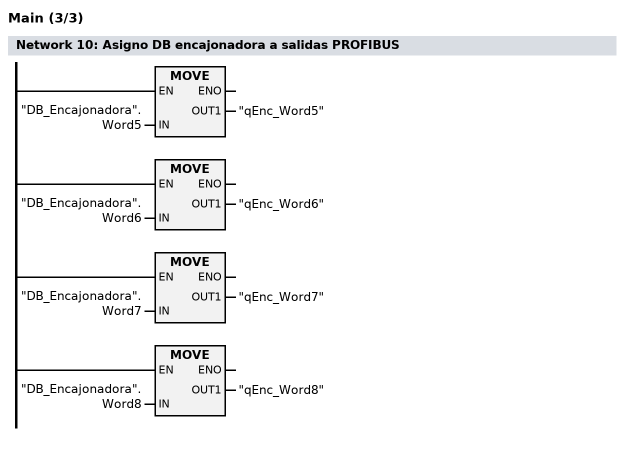
   RUNG wire#powerrail
      Move(in := "DB_Encajonadora".Word5, out1 => "qEnc_Word5")
   END_RUNG
   RUNG wire#powerrail
      Move(in := "DB_Encajonadora".Word6, out1 => "qEnc_Word6")
   END_RUNG
   RUNG wire#powerrail
      Move(in := "DB_Encajonadora".Word7, out1 => "qEnc_Word7")
   END_RUNG
   RUNG wire#powerrail
      Move(in := "DB_Encajonadora".Word8, out1 => "qEnc_Word8")
   END_RUNG
   // the same network as SCL:
   "qEnc_Word5" := "DB_Encajonadora".Word5;
   "qEnc_Word6" := "DB_Encajonadora".Word6;
   "qEnc_Word7" := "DB_Encajonadora".Word7;
   "qEnc_Word8" := "DB_Encajonadora".Word8;
END_REGION
END_ORGANIZATION_BLOCK

ORGANIZATION_BLOCK "Cyclic interrupt"   // OB30, LAD, CyclicInterrupt
{ S7_Optimized_Access := 'TRUE' }
VERSION : 0.1
   VAR_INPUT
      Initial_Call : Bool;   // Initial call of this OB
      Event_Count : Int;   // Events discarded
   END_VAR
BEGIN

REGION Network 1: Move
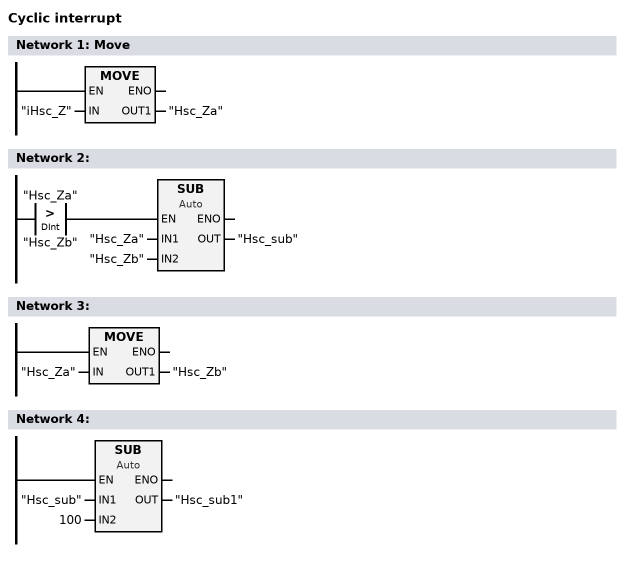
   RUNG wire#powerrail
      Move(in := "iHsc_Z", out1 => "Hsc_Za")
   END_RUNG
   // the same network as SCL:
   "Hsc_Za" := "iHsc_Z";
END_REGION

REGION Network 2
   RUNG wire#powerrail
      { S7_Templates := "SrcType := DInt" } GT_Contact(in1 := "Hsc_Za", in2 := "Hsc_Zb")
      Sub(in1 := "Hsc_Za", in2 := "Hsc_Zb", out => "Hsc_sub")
   END_RUNG
   // the same network as SCL:
   IF "Hsc_Za" > "Hsc_Zb" THEN "Hsc_sub" := "Hsc_Za" - "Hsc_Zb"; END_IF;
END_REGION

REGION Network 3
   RUNG wire#powerrail
      Move(in := "Hsc_Za", out1 => "Hsc_Zb")
   END_RUNG
   // the same network as SCL:
   "Hsc_Zb" := "Hsc_Za";
END_REGION

REGION Network 4
   RUNG wire#powerrail
      Sub(in1 := "Hsc_sub", in2 := 100, out => "Hsc_sub1")
   END_RUNG
   // the same network as SCL:
   "Hsc_sub1" := "Hsc_sub" - 100;
END_REGION
END_ORGANIZATION_BLOCK

// folder: ESTANDAR

FUNCTION_BLOCK "Motor M&CM"   // FB2, LAD
TITLE = Motor Marcha & Contra-Marcha
{ S7_Optimized_Access := 'TRUE' }
VERSION : 0.1
   VAR_INPUT
      iOrdMar_Dir : Bool;
      iOrdMar_Rev : Bool;
      iConfMar_Dir : Bool;
      iConfMar_Rev : Bool;
      iGMT : Bool;
      iTConf_Warn : Time;
      iTConf_Fall : Time;
      iTRearranque : Time;
   END_VAR
   VAR_OUTPUT
      oMar_Dir : Bool;
      oMar_Rev : Bool;
      oWarning_CTC_Dir : Bool;
      oWarning_CTC_Rev : Bool;
      oFall_CTC_Dir : Bool;
      oFall_CTC_Rev : Bool;
      oFall_GMT : Bool;
   END_VAR
   VAR
      IEC_Timer_0_Instance : IEC_TIMER;
      IEC_Timer_0_Instance_1 : IEC_TIMER;
      IEC_Timer_0_Instance_2 : IEC_TIMER;
      IEC_Timer_0_Instance_3 : IEC_TIMER;
      IEC_Timer_0_Instance_4 : IEC_TIMER;
      MarDir_Aux : Bool;
      MarRev_Aux : Bool;
   END_VAR
   VAR_TEMP
      Fall_GMT_Aux : Bool;
      Fall_CTC_Dir_Aux : Bool;
      Fall_CTC_Rev_Aux : Bool;
      Habil_Mov : Bool;
   END_VAR
   VAR_TEMP   // added for the SCL form of the ladder/FBD networks
      _w1 : Bool;
   END_VAR
BEGIN

REGION Network 1: Falla Guardamotor
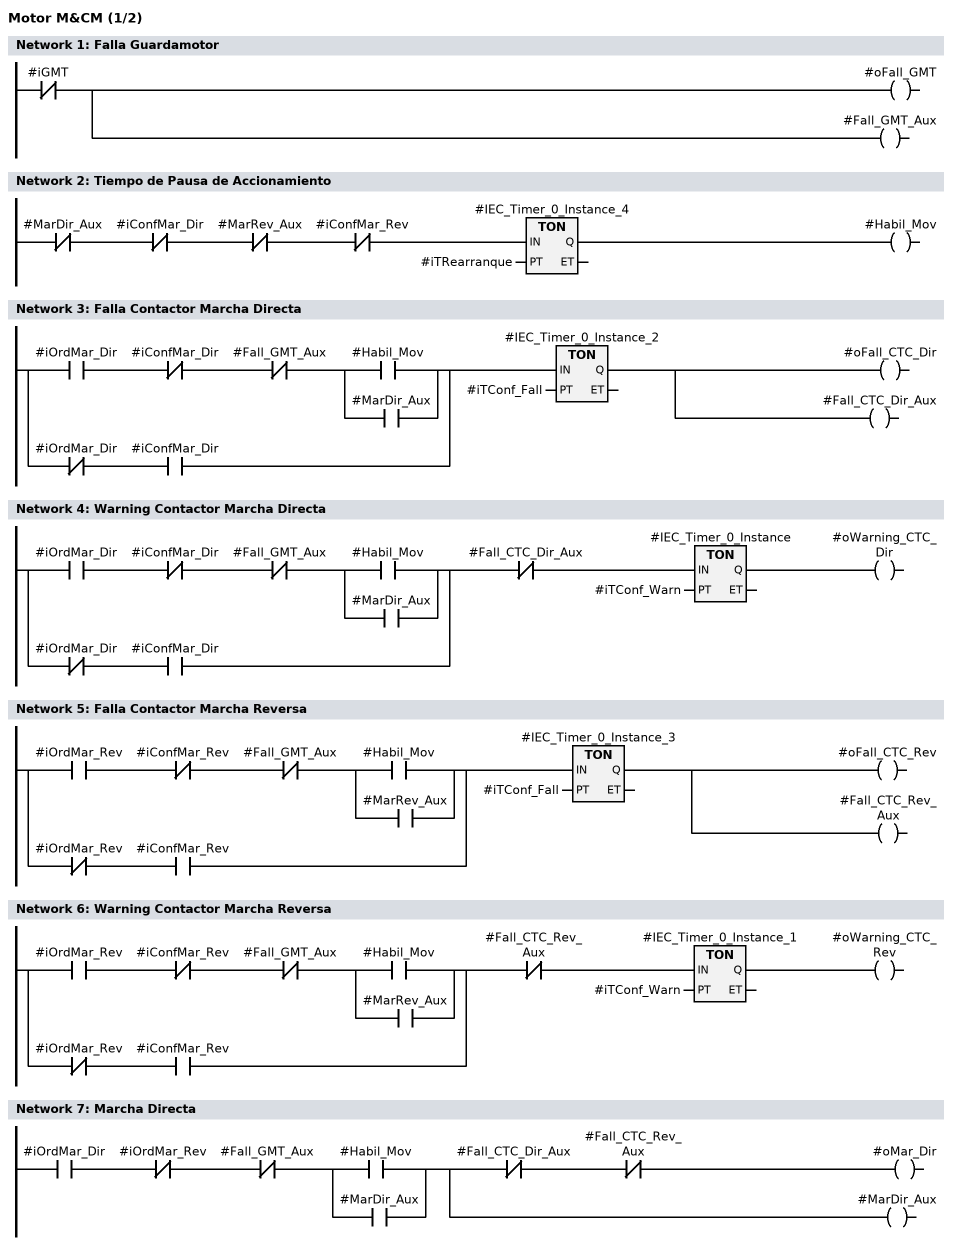
   RUNG wire#powerrail
      I_Contact( #iGMT )
      wire#w1
      Coil( #oFall_GMT )
   END_RUNG
   RUNG wire#w1
      Coil( #Fall_GMT_Aux )
   END_RUNG
   // the same network as SCL:
   #oFall_GMT := NOT #iGMT;
   #Fall_GMT_Aux := NOT #iGMT;
END_REGION

REGION Network 2: Tiempo de Pausa de Accionamiento
   #IEC_Timer_0_Instance_4.TON(IN := NOT #MarDir_Aux AND NOT #iConfMar_Dir AND NOT #MarRev_Aux AND NOT #iConfMar_Rev,
                           PT := #iTRearranque);
   #Habil_Mov := #IEC_Timer_0_Instance_4.Q;
END_REGION

REGION Network 3: Falla Contactor Marcha Directa
   #IEC_Timer_0_Instance_2.TON(IN := (#iOrdMar_Dir AND NOT #iConfMar_Dir AND NOT #Fall_GMT_Aux AND (#Habil_Mov OR #MarDir_Aux)) OR (NOT #iOrdMar_Dir AND #iConfMar_Dir),
                           PT := #iTConf_Fall);
   #oFall_CTC_Dir := #IEC_Timer_0_Instance_2.Q;
   #Fall_CTC_Dir_Aux := #IEC_Timer_0_Instance_2.Q;
END_REGION

REGION Network 4: Warning Contactor Marcha Directa
   #IEC_Timer_0_Instance.TON(IN := ((#iOrdMar_Dir AND NOT #iConfMar_Dir AND NOT #Fall_GMT_Aux AND (#Habil_Mov OR #MarDir_Aux)) OR (NOT #iOrdMar_Dir AND #iConfMar_Dir)) AND NOT #Fall_CTC_Dir_Aux,
                           PT := #iTConf_Warn);
   #oWarning_CTC_Dir := #IEC_Timer_0_Instance.Q;
END_REGION

REGION Network 5: Falla Contactor Marcha Reversa
   #IEC_Timer_0_Instance_3.TON(IN := (#iOrdMar_Rev AND NOT #iConfMar_Rev AND NOT #Fall_GMT_Aux AND (#Habil_Mov OR #MarRev_Aux)) OR (NOT #iOrdMar_Rev AND #iConfMar_Rev),
                           PT := #iTConf_Fall);
   #oFall_CTC_Rev := #IEC_Timer_0_Instance_3.Q;
   #Fall_CTC_Rev_Aux := #IEC_Timer_0_Instance_3.Q;
END_REGION

REGION Network 6: Warning Contactor Marcha Reversa
   #IEC_Timer_0_Instance_1.TON(IN := ((#iOrdMar_Rev AND NOT #iConfMar_Rev AND NOT #Fall_GMT_Aux AND (#Habil_Mov OR #MarRev_Aux)) OR (NOT #iOrdMar_Rev AND #iConfMar_Rev)) AND NOT #Fall_CTC_Rev_Aux,
                           PT := #iTConf_Warn);
   #oWarning_CTC_Rev := #IEC_Timer_0_Instance_1.Q;
END_REGION

REGION Network 7: Marcha Directa
   RUNG wire#powerrail
      Contact( #iOrdMar_Dir )
      I_Contact( #iOrdMar_Rev )
      I_Contact( #Fall_GMT_Aux )
      wire#w1
      Contact( #Habil_Mov )
      wire#w2
      I_Contact( #Fall_CTC_Dir_Aux )
      I_Contact( #Fall_CTC_Rev_Aux )
      Coil( #oMar_Dir )
   END_RUNG
   RUNG wire#w1
      Contact( #MarDir_Aux )
   END_RUNG wire#w2
   RUNG wire#w2
      Coil( #MarDir_Aux )
   END_RUNG
   // the same network as SCL:
   #_w1 := #iOrdMar_Dir AND NOT #iOrdMar_Rev AND NOT #Fall_GMT_Aux AND (#Habil_Mov OR #MarDir_Aux);
   #oMar_Dir := #_w1 AND NOT #Fall_CTC_Dir_Aux AND NOT #Fall_CTC_Rev_Aux;
   #MarDir_Aux := #_w1;
END_REGION

REGION Network 8: Marcha Reversa
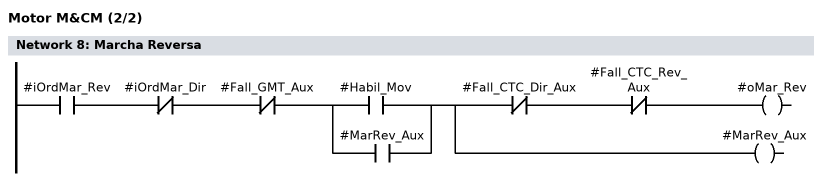
   RUNG wire#powerrail
      Contact( #iOrdMar_Rev )
      I_Contact( #iOrdMar_Dir )
      I_Contact( #Fall_GMT_Aux )
      wire#w1
      Contact( #Habil_Mov )
      wire#w2
      I_Contact( #Fall_CTC_Dir_Aux )
      I_Contact( #Fall_CTC_Rev_Aux )
      Coil( #oMar_Rev )
   END_RUNG
   RUNG wire#w1
      Contact( #MarRev_Aux )
   END_RUNG wire#w2
   RUNG wire#w2
      Coil( #MarRev_Aux )
   END_RUNG
   // the same network as SCL:
   #_w1 := #iOrdMar_Rev AND NOT #iOrdMar_Dir AND NOT #Fall_GMT_Aux AND (#Habil_Mov OR #MarRev_Aux);
   #oMar_Rev := #_w1 AND NOT #Fall_CTC_Dir_Aux AND NOT #Fall_CTC_Rev_Aux;
   #MarRev_Aux := #_w1;
END_REGION
END_FUNCTION_BLOCK

FUNCTION_BLOCK "FB_VAR_MOT"   // FB4, LAD
{ S7_Optimized_Access := 'FALSE' }
VERSION : 0.1
   VAR_INPUT
      "CMD Mar Dir" : Bool;   // Comando Marcha Directa
      "CMD Mar Rev" : Bool;   // Comando Marcha Reversa
      "HAB  Mar" : Bool;   // Habilita Marcha
      "SP Vel" : Real;   // Setpoint de Velocidad
      Reset : Bool;   // Comando resetear falla
      Fault : Bool;   // Indica variador en falla
      Ready : Bool;   // Indica variador Ready
      Ton_Freno : Time := T#400ms;
      Ton_Mar : Time := T#100ms;
      Tof_Freno : Time := T#100ms;
      Tof_Mar : Time := T#200ms;
   END_VAR
   VAR_OUTPUT
      Marcha : Bool;   // Orden de marcha a variador
      "Inv Giro" : Bool;   // Orden de invertir sentido de giro a variador
      "Reset Fault" : Bool;   // Reset Fault a variador
      Velocidad : Word;   // Referencia de Velocidad a variador
      Freno : Bool;   // Apertura de Freno
      Falla : Bool;   // Indica falla del variador
      Warning : Bool;   // Indica variador no Ready
   END_VAR
   VAR
      IEC_Timer_Freno : TON_TIME;
      IEC_Timer_Motor : TON_TIME;
      IEC_Timer_Reset : TOF_TIME;
      "_CMD Marcha Dir" : Bool;
      "_CMD Marcha Rev" : Bool;
      _CMD_AbrirFreno : Bool;
      IEC_Timer_0_Instance : TON_TIME;
      IEC_Timer_0_Instance_1 : TOF_TIME;
      IEC_Timer_0_Instance_2 : TOF_TIME;
      Ord_Marcha : Bool;
      Mem_Inv : Bool;
   END_VAR
   VAR_TEMP
      Vel_Real : Real;
      Vel_Int : Int;
      _Hab_Abrir_Freno : Bool;
      "Pre Marcha" : Bool;
      Aux : Bool;
      Freno_Aux : Bool;
   END_VAR
   VAR_TEMP   // added for the SCL form of the ladder/FBD networks
      _w1 : Bool;
      _w2 : Bool;
      _w3 : Bool;
   END_VAR
BEGIN

REGION Network 1: #Aux
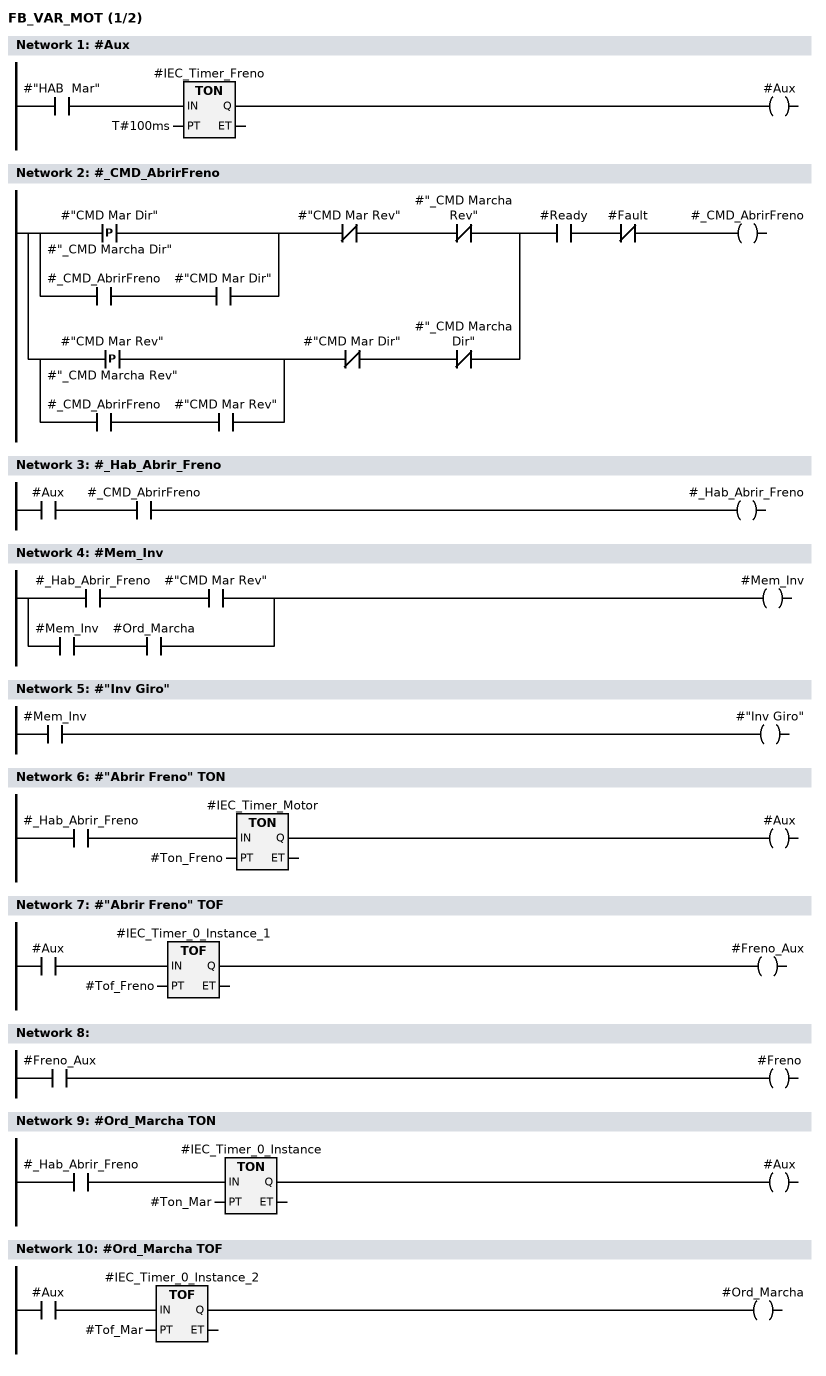
   #IEC_Timer_Freno(IN := #"HAB  Mar", PT := T#100ms);   // TON
   #Aux := #IEC_Timer_Freno.Q;
END_REGION

REGION Network 2: #_CMD_AbrirFreno
   RUNG wire#powerrail
      P_Contact(operand := #"CMD Mar Dir", bit := #"_CMD Marcha Dir")
      wire#w1
      I_Contact( #"CMD Mar Rev" )
      I_Contact( #"_CMD Marcha Rev" )
      wire#w2
      Contact( #Ready )
      I_Contact( #Fault )
      Coil( #_CMD_AbrirFreno )
   END_RUNG
   RUNG wire#powerrail
      Contact( #_CMD_AbrirFreno )
      Contact( #"CMD Mar Dir" )
   END_RUNG wire#w1
   RUNG wire#powerrail
      P_Contact(operand := #"CMD Mar Rev", bit := #"_CMD Marcha Rev")
      wire#w3
      I_Contact( #"CMD Mar Dir" )
      I_Contact( #"_CMD Marcha Dir" )
   END_RUNG wire#w2
   RUNG wire#powerrail
      Contact( #_CMD_AbrirFreno )
      Contact( #"CMD Mar Rev" )
   END_RUNG wire#w3
   // the same network as SCL:
   #_w1 := #"CMD Mar Dir" AND NOT #"_CMD Marcha Dir";   // rising edge of #"CMD Mar Dir"
   #"_CMD Marcha Dir" := #"CMD Mar Dir";
   #_w3 := (#_w1 OR (#_CMD_AbrirFreno AND #"CMD Mar Dir")) AND NOT #"CMD Mar Rev" AND NOT #"_CMD Marcha Rev";
   #_w2 := #"CMD Mar Rev" AND NOT #"_CMD Marcha Rev";   // rising edge of #"CMD Mar Rev"
   #"_CMD Marcha Rev" := #"CMD Mar Rev";
   #_CMD_AbrirFreno := (#_w3 OR ((#_w2 OR (#_CMD_AbrirFreno AND #"CMD Mar Rev")) AND NOT #"CMD Mar Dir" AND NOT #"_CMD Marcha Dir")) AND #Ready AND NOT #Fault;
END_REGION

REGION Network 3: #_Hab_Abrir_Freno
   RUNG wire#powerrail
      Contact( #Aux )
      Contact( #_CMD_AbrirFreno )
      Coil( #_Hab_Abrir_Freno )
   END_RUNG
   // the same network as SCL:
   #_Hab_Abrir_Freno := #Aux AND #_CMD_AbrirFreno;
END_REGION

REGION Network 4: #Mem_Inv
   RUNG wire#powerrail
      Contact( #_Hab_Abrir_Freno )
      Contact( #"CMD Mar Rev" )
      wire#w1
      Coil( #Mem_Inv )
   END_RUNG
   RUNG wire#powerrail
      Contact( #Mem_Inv )
      Contact( #Ord_Marcha )
   END_RUNG wire#w1
   // the same network as SCL:
   #Mem_Inv := (#_Hab_Abrir_Freno AND #"CMD Mar Rev") OR (#Mem_Inv AND #Ord_Marcha);
END_REGION

REGION Network 5: #"Inv Giro"
   RUNG wire#powerrail
      Contact( #Mem_Inv )
      Coil( #"Inv Giro" )
   END_RUNG
   // the same network as SCL:
   #"Inv Giro" := #Mem_Inv;
END_REGION

REGION Network 6: #"Abrir Freno" TON
   #IEC_Timer_Motor(IN := #_Hab_Abrir_Freno, PT := #Ton_Freno);   // TON
   #Aux := #IEC_Timer_Motor.Q;
END_REGION

REGION Network 7: #"Abrir Freno" TOF
   #IEC_Timer_0_Instance_1(IN := #Aux, PT := #Tof_Freno);   // TOF
   #Freno_Aux := #IEC_Timer_0_Instance_1.Q;
END_REGION

REGION Network 8
   RUNG wire#powerrail
      Contact( #Freno_Aux )
      Coil( #Freno )
   END_RUNG
   // the same network as SCL:
   #Freno := #Freno_Aux;
END_REGION

REGION Network 9: #Ord_Marcha TON
   #IEC_Timer_0_Instance(IN := #_Hab_Abrir_Freno, PT := #Ton_Mar);   // TON
   #Aux := #IEC_Timer_0_Instance.Q;
END_REGION

REGION Network 10: #Ord_Marcha TOF
   #IEC_Timer_0_Instance_2(IN := #Aux, PT := #Tof_Mar);   // TOF
   #Ord_Marcha := #IEC_Timer_0_Instance_2.Q;
END_REGION

REGION Network 11: #Marcha
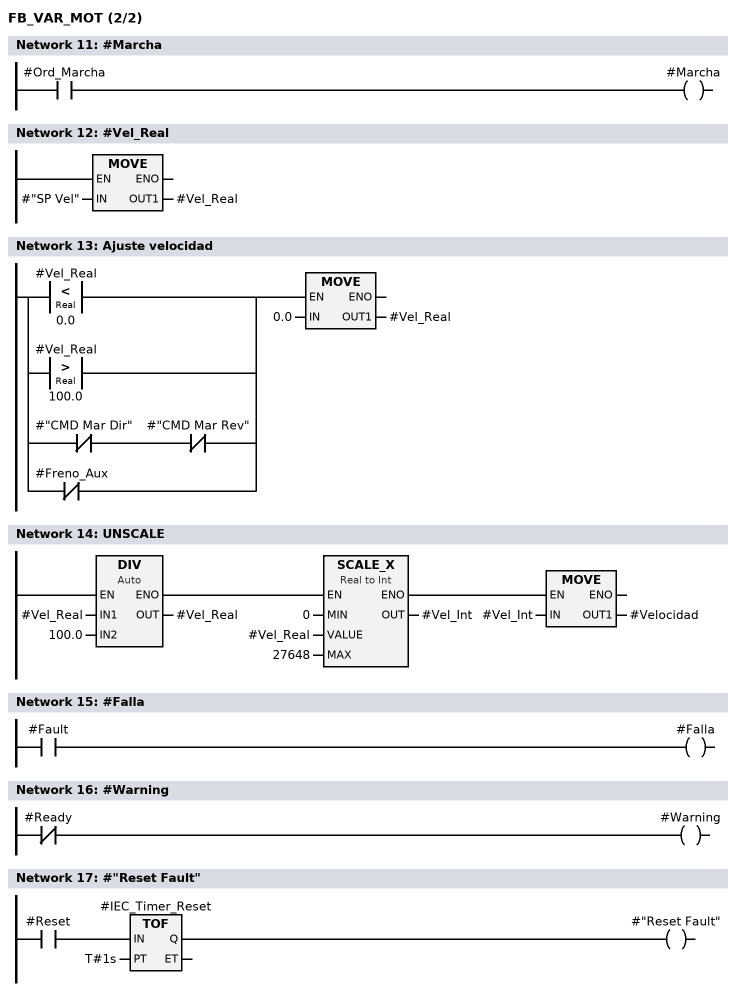
   RUNG wire#powerrail
      Contact( #Ord_Marcha )
      Coil( #Marcha )
   END_RUNG
   // the same network as SCL:
   #Marcha := #Ord_Marcha;
END_REGION

REGION Network 12: #Vel_Real
   RUNG wire#powerrail
      { S7_GenerateENO := "TRUE" } Move(in := #"SP Vel", out1 => #Vel_Real)
   END_RUNG
   // the same network as SCL:
   #Vel_Real := #"SP Vel";
END_REGION

REGION Network 13: Ajuste velocidad
   RUNG wire#powerrail
      { S7_Templates := "SrcType := Real" } LT_Contact(in1 := #Vel_Real, in2 := 0.0)
      wire#w1
      { S7_GenerateENO := "TRUE" } Move(in := 0.0, out1 => #Vel_Real)
   END_RUNG
   RUNG wire#powerrail
      { S7_Templates := "SrcType := Real" } GT_Contact(in1 := #Vel_Real, in2 := 100.0)
   END_RUNG wire#w1
   RUNG wire#powerrail
      I_Contact( #"CMD Mar Dir" )
      I_Contact( #"CMD Mar Rev" )
   END_RUNG wire#w1
   RUNG wire#powerrail
      I_Contact( #Freno_Aux )
   END_RUNG wire#w1
   // the same network as SCL:
   IF (#Vel_Real < 0.0) OR (#Vel_Real > 100.0) OR (NOT #"CMD Mar Dir" AND NOT #"CMD Mar Rev") OR NOT #Freno_Aux THEN
       #Vel_Real := 0.0;
   END_IF;
END_REGION

REGION Network 14: UNSCALE
   RUNG wire#powerrail
      Div(in1 := #Vel_Real, in2 := 100.0, out => #Vel_Real)
      { S7_Templates := "[SrcType := Real, DestType := Int]" } Scale(min := 0, value := #Vel_Real, max := 27648, out => #Vel_Int)
      { S7_GenerateENO := "TRUE" } Move(in := #Vel_Int, out1 => #Velocidad)
   END_RUNG
   // the same network as SCL:
   #Vel_Real := #Vel_Real / 100.0;
   #Vel_Int := SCALE_X(MIN := 0, VALUE := #Vel_Real, MAX := 27648);
   #Velocidad := #Vel_Int;
END_REGION

REGION Network 15: #Falla
   RUNG wire#powerrail
      Contact( #Fault )
      Coil( #Falla )
   END_RUNG
   // the same network as SCL:
   #Falla := #Fault;
END_REGION

REGION Network 16: #Warning
   RUNG wire#powerrail
      I_Contact( #Ready )
      Coil( #Warning )
   END_RUNG
   // the same network as SCL:
   #Warning := NOT #Ready;
END_REGION

REGION Network 17: #"Reset Fault"
   #IEC_Timer_Reset(IN := #Reset, PT := T#1s);   // TOF
   #"Reset Fault" := #IEC_Timer_Reset.Q;
END_REGION
END_FUNCTION_BLOCK

FUNCTION_BLOCK "Motor Simple"   // FB5, LAD
{ S7_Optimized_Access := 'TRUE' }
VERSION : 0.1
   VAR_INPUT
      iOrdMar : Bool;
      iConfMar : Bool;
      iGMT : Bool;
      iTConf_Warn : Time;
      iTConf_Fall : Time;
      iTRearranque : Time;
   END_VAR
   VAR_OUTPUT
      oMarcha : Bool;
      oWarning_CTC : Bool;
      oFall_CTC : Bool;
      oFall_GMT : Bool;
   END_VAR
   VAR
      IEC_Timer_0_Instance : IEC_TIMER;
      IEC_Timer_0_Instance_1 : IEC_TIMER;
      IEC_Timer_0_Instance_2 : IEC_TIMER;
      Mar_Aux : Bool;
   END_VAR
   VAR_TEMP
      Fall_GMT_Aux : Bool;
      Fall_CTC_Aux : Bool;
      Habil_Mov : Bool;
   END_VAR
BEGIN

REGION Network 1: Falla Guardamotor
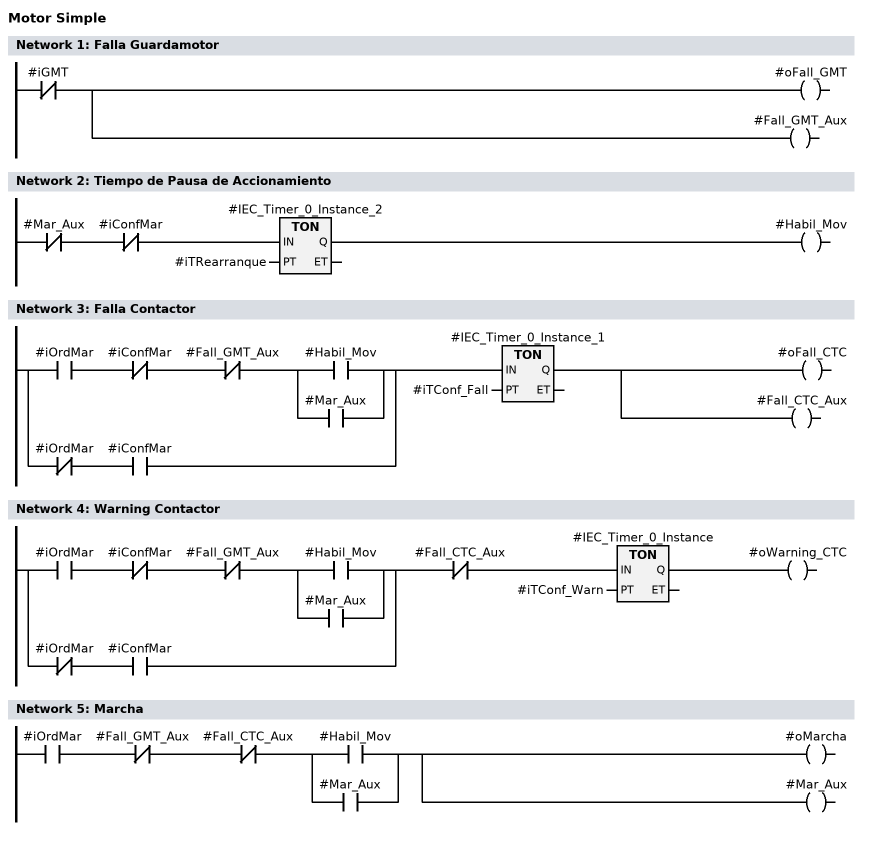
   RUNG wire#powerrail
      I_Contact( #iGMT )
      wire#w1
      Coil( #oFall_GMT )
   END_RUNG
   RUNG wire#w1
      Coil( #Fall_GMT_Aux )
   END_RUNG
   // the same network as SCL:
   #oFall_GMT := NOT #iGMT;
   #Fall_GMT_Aux := NOT #iGMT;
END_REGION

REGION Network 2: Tiempo de Pausa de Accionamiento
   #IEC_Timer_0_Instance_2.TON(IN := NOT #Mar_Aux AND NOT #iConfMar, PT := #iTRearranque);
   #Habil_Mov := #IEC_Timer_0_Instance_2.Q;
END_REGION

REGION Network 3: Falla Contactor
   #IEC_Timer_0_Instance_1.TON(IN := (#iOrdMar AND NOT #iConfMar AND NOT #Fall_GMT_Aux AND (#Habil_Mov OR #Mar_Aux)) OR (NOT #iOrdMar AND #iConfMar),
                           PT := #iTConf_Fall);
   #oFall_CTC := #IEC_Timer_0_Instance_1.Q;
   #Fall_CTC_Aux := #IEC_Timer_0_Instance_1.Q;
END_REGION

REGION Network 4: Warning Contactor
   #IEC_Timer_0_Instance.TON(IN := ((#iOrdMar AND NOT #iConfMar AND NOT #Fall_GMT_Aux AND (#Habil_Mov OR #Mar_Aux)) OR (NOT #iOrdMar AND #iConfMar)) AND NOT #Fall_CTC_Aux,
                           PT := #iTConf_Warn);
   #oWarning_CTC := #IEC_Timer_0_Instance.Q;
END_REGION

REGION Network 5: Marcha
   RUNG wire#powerrail
      Contact( #iOrdMar )
      I_Contact( #Fall_GMT_Aux )
      I_Contact( #Fall_CTC_Aux )
      wire#w1
      Contact( #Habil_Mov )
      wire#w2
      Coil( #oMarcha )
   END_RUNG
   RUNG wire#w1
      Contact( #Mar_Aux )
   END_RUNG wire#w2
   RUNG wire#w2
      Coil( #Mar_Aux )
   END_RUNG
   // the same network as SCL:
   #oMarcha := #iOrdMar AND NOT #Fall_GMT_Aux AND NOT #Fall_CTC_Aux AND (#Habil_Mov OR #Mar_Aux);
   #Mar_Aux := #oMarcha;
END_REGION
END_FUNCTION_BLOCK

FUNCTION_BLOCK "FB_VLV_2_POS"   // FB6, LAD
{ S7_Optimized_Access := 'FALSE' }